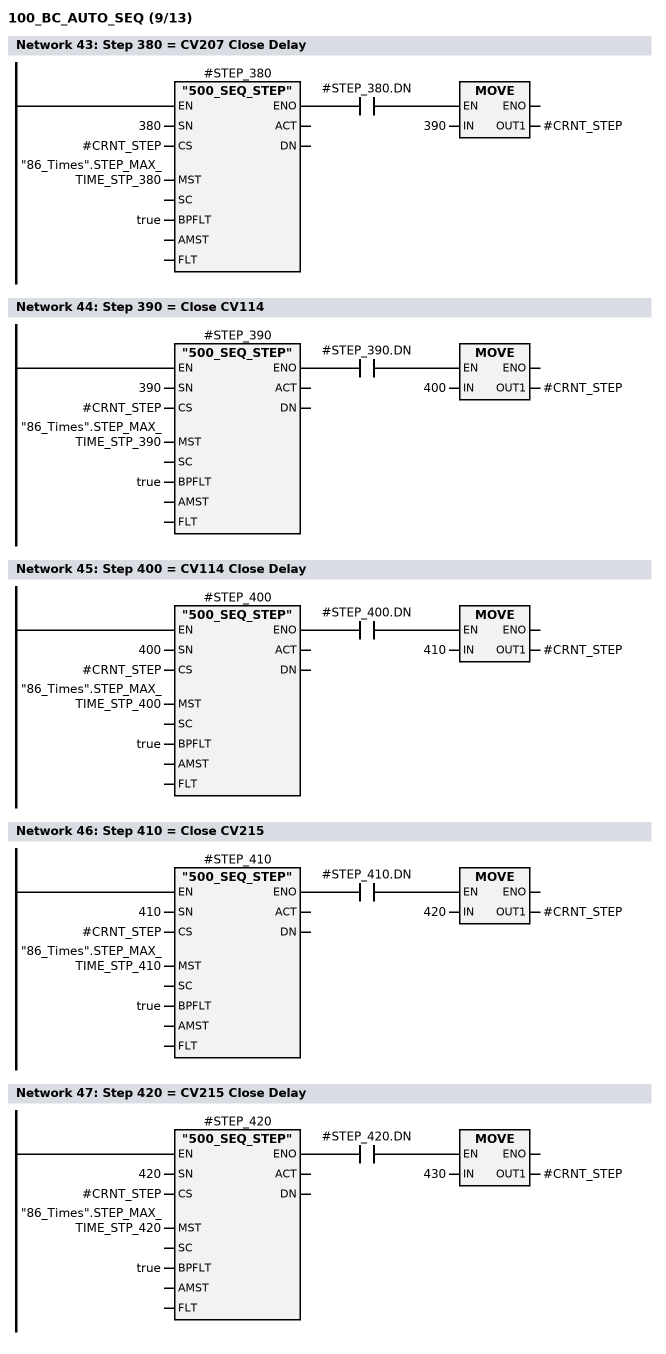
   RUNG wire#powerrail
      #STEP_380(SN := 380, CS := #CRNT_STEP, MST := "86_Times".STEP_MAX_TIME_STP_380, SC :=, BPFLT := true, AMST :=, FLT :=, ACT =>, DN =>)
      Contact( #STEP_380.DN )
      Move(in := 390, out1 => #CRNT_STEP)
   END_RUNG
   // the same network as SCL:
   #STEP_380(SN := 380, CS := #CRNT_STEP, MST := "86_Times".STEP_MAX_TIME_STP_380, BPFLT := true, ENO => #_w1);   // "500_SEQ_STEP"
   IF #_w1 AND #STEP_380.DN THEN #CRNT_STEP := 390; END_IF;
END_REGION

REGION Network 44: Step 390 = Close CV114
   RUNG wire#powerrail
      #STEP_390(SN := 390, CS := #CRNT_STEP, MST := "86_Times".STEP_MAX_TIME_STP_390, SC :=, BPFLT := true, AMST :=, FLT :=, ACT =>, DN =>)
      Contact( #STEP_390.DN )
      Move(in := 400, out1 => #CRNT_STEP)
   END_RUNG
   // the same network as SCL:
   #STEP_390(SN := 390, CS := #CRNT_STEP, MST := "86_Times".STEP_MAX_TIME_STP_390, BPFLT := true, ENO => #_w1);   // "500_SEQ_STEP"
   IF #_w1 AND #STEP_390.DN THEN #CRNT_STEP := 400; END_IF;
END_REGION

REGION Network 45: Step 400 = CV114 Close Delay
   RUNG wire#powerrail
      #STEP_400(SN := 400, CS := #CRNT_STEP, MST := "86_Times".STEP_MAX_TIME_STP_400, SC :=, BPFLT := true, AMST :=, FLT :=, ACT =>, DN =>)
      Contact( #STEP_400.DN )
      Move(in := 410, out1 => #CRNT_STEP)
   END_RUNG
   // the same network as SCL:
   #STEP_400(SN := 400, CS := #CRNT_STEP, MST := "86_Times".STEP_MAX_TIME_STP_400, BPFLT := true, ENO => #_w1);   // "500_SEQ_STEP"
   IF #_w1 AND #STEP_400.DN THEN #CRNT_STEP := 410; END_IF;
END_REGION

REGION Network 46: Step 410 = Close CV215
   RUNG wire#powerrail
      #STEP_410(SN := 410, CS := #CRNT_STEP, MST := "86_Times".STEP_MAX_TIME_STP_410, SC :=, BPFLT := true, AMST :=, FLT :=, ACT =>, DN =>)
      Contact( #STEP_410.DN )
      Move(in := 420, out1 => #CRNT_STEP)
   END_RUNG
   // the same network as SCL:
   #STEP_410(SN := 410, CS := #CRNT_STEP, MST := "86_Times".STEP_MAX_TIME_STP_410, BPFLT := true, ENO => #_w1);   // "500_SEQ_STEP"
   IF #_w1 AND #STEP_410.DN THEN #CRNT_STEP := 420; END_IF;
END_REGION

REGION Network 47: Step 420 = CV215 Close Delay
   RUNG wire#powerrail
      #STEP_420(SN := 420, CS := #CRNT_STEP, MST := "86_Times".STEP_MAX_TIME_STP_420, SC :=, BPFLT := true, AMST :=, FLT :=, ACT =>, DN =>)
      Contact( #STEP_420.DN )
      Move(in := 430, out1 => #CRNT_STEP)
   END_RUNG
   // the same network as SCL:
   #STEP_420(SN := 420, CS := #CRNT_STEP, MST := "86_Times".STEP_MAX_TIME_STP_420, BPFLT := true, ENO => #_w1);   // "500_SEQ_STEP"
   IF #_w1 AND #STEP_420.DN THEN #CRNT_STEP := 430; END_IF;
END_REGION

REGION Network 48: Step 430 = Close CV216
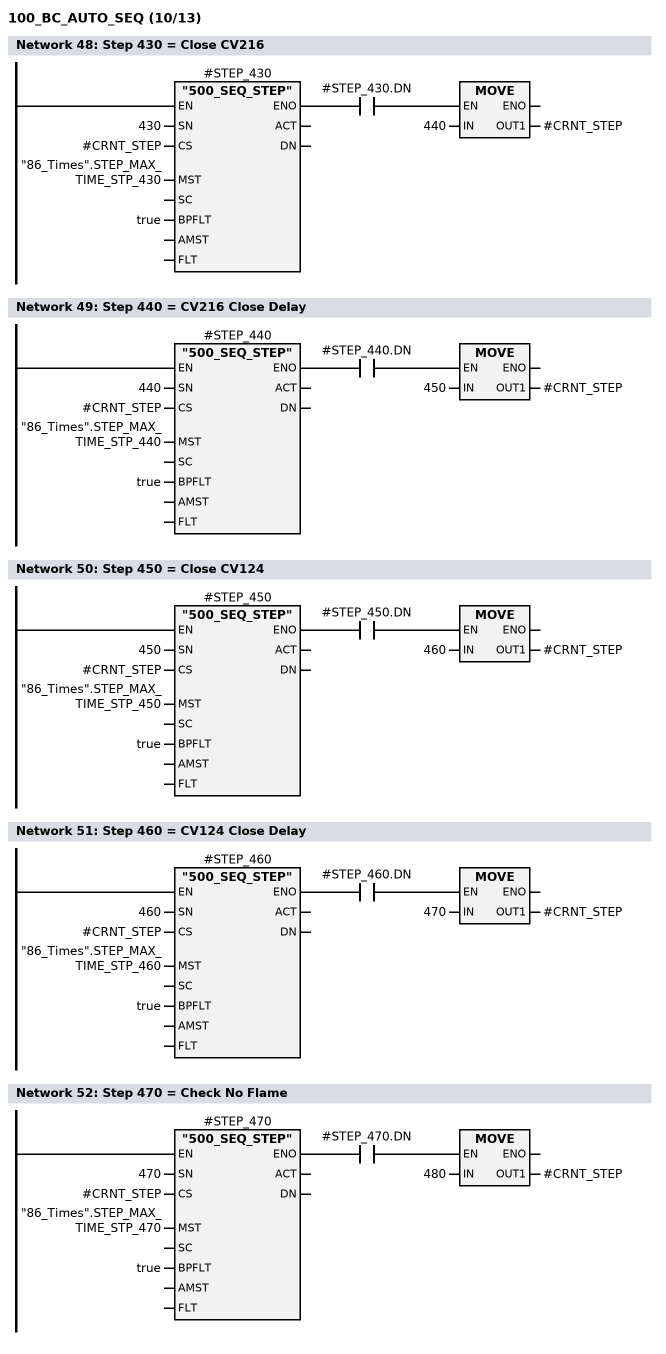
   RUNG wire#powerrail
      #STEP_430(SN := 430, CS := #CRNT_STEP, MST := "86_Times".STEP_MAX_TIME_STP_430, SC :=, BPFLT := true, AMST :=, FLT :=, ACT =>, DN =>)
      Contact( #STEP_430.DN )
      Move(in := 440, out1 => #CRNT_STEP)
   END_RUNG
   // the same network as SCL:
   #STEP_430(SN := 430, CS := #CRNT_STEP, MST := "86_Times".STEP_MAX_TIME_STP_430, BPFLT := true, ENO => #_w1);   // "500_SEQ_STEP"
   IF #_w1 AND #STEP_430.DN THEN #CRNT_STEP := 440; END_IF;
END_REGION

REGION Network 49: Step 440 = CV216 Close Delay
   RUNG wire#powerrail
      #STEP_440(SN := 440, CS := #CRNT_STEP, MST := "86_Times".STEP_MAX_TIME_STP_440, SC :=, BPFLT := true, AMST :=, FLT :=, ACT =>, DN =>)
      Contact( #STEP_440.DN )
      Move(in := 450, out1 => #CRNT_STEP)
   END_RUNG
   // the same network as SCL:
   #STEP_440(SN := 440, CS := #CRNT_STEP, MST := "86_Times".STEP_MAX_TIME_STP_440, BPFLT := true, ENO => #_w1);   // "500_SEQ_STEP"
   IF #_w1 AND #STEP_440.DN THEN #CRNT_STEP := 450; END_IF;
END_REGION

REGION Network 50: Step 450 = Close CV124
   RUNG wire#powerrail
      #STEP_450(SN := 450, CS := #CRNT_STEP, MST := "86_Times".STEP_MAX_TIME_STP_450, SC :=, BPFLT := true, AMST :=, FLT :=, ACT =>, DN =>)
      Contact( #STEP_450.DN )
      Move(in := 460, out1 => #CRNT_STEP)
   END_RUNG
   // the same network as SCL:
   #STEP_450(SN := 450, CS := #CRNT_STEP, MST := "86_Times".STEP_MAX_TIME_STP_450, BPFLT := true, ENO => #_w1);   // "500_SEQ_STEP"
   IF #_w1 AND #STEP_450.DN THEN #CRNT_STEP := 460; END_IF;
END_REGION

REGION Network 51: Step 460 = CV124 Close Delay
   RUNG wire#powerrail
      #STEP_460(SN := 460, CS := #CRNT_STEP, MST := "86_Times".STEP_MAX_TIME_STP_460, SC :=, BPFLT := true, AMST :=, FLT :=, ACT =>, DN =>)
      Contact( #STEP_460.DN )
      Move(in := 470, out1 => #CRNT_STEP)
   END_RUNG
   // the same network as SCL:
   #STEP_460(SN := 460, CS := #CRNT_STEP, MST := "86_Times".STEP_MAX_TIME_STP_460, BPFLT := true, ENO => #_w1);   // "500_SEQ_STEP"
   IF #_w1 AND #STEP_460.DN THEN #CRNT_STEP := 470; END_IF;
END_REGION

REGION Network 52: Step 470 = Check No Flame
   RUNG wire#powerrail
      #STEP_470(SN := 470, CS := #CRNT_STEP, MST := "86_Times".STEP_MAX_TIME_STP_470, SC :=, BPFLT := true, AMST :=, FLT :=, ACT =>, DN =>)
      Contact( #STEP_470.DN )
      Move(in := 480, out1 => #CRNT_STEP)
   END_RUNG
   // the same network as SCL:
   #STEP_470(SN := 470, CS := #CRNT_STEP, MST := "86_Times".STEP_MAX_TIME_STP_470, BPFLT := true, ENO => #_w1);   // "500_SEQ_STEP"
   IF #_w1 AND #STEP_470.DN THEN #CRNT_STEP := 480; END_IF;
END_REGION

REGION Network 53: Step 480 = Burn Stopped Confirmation To IGG
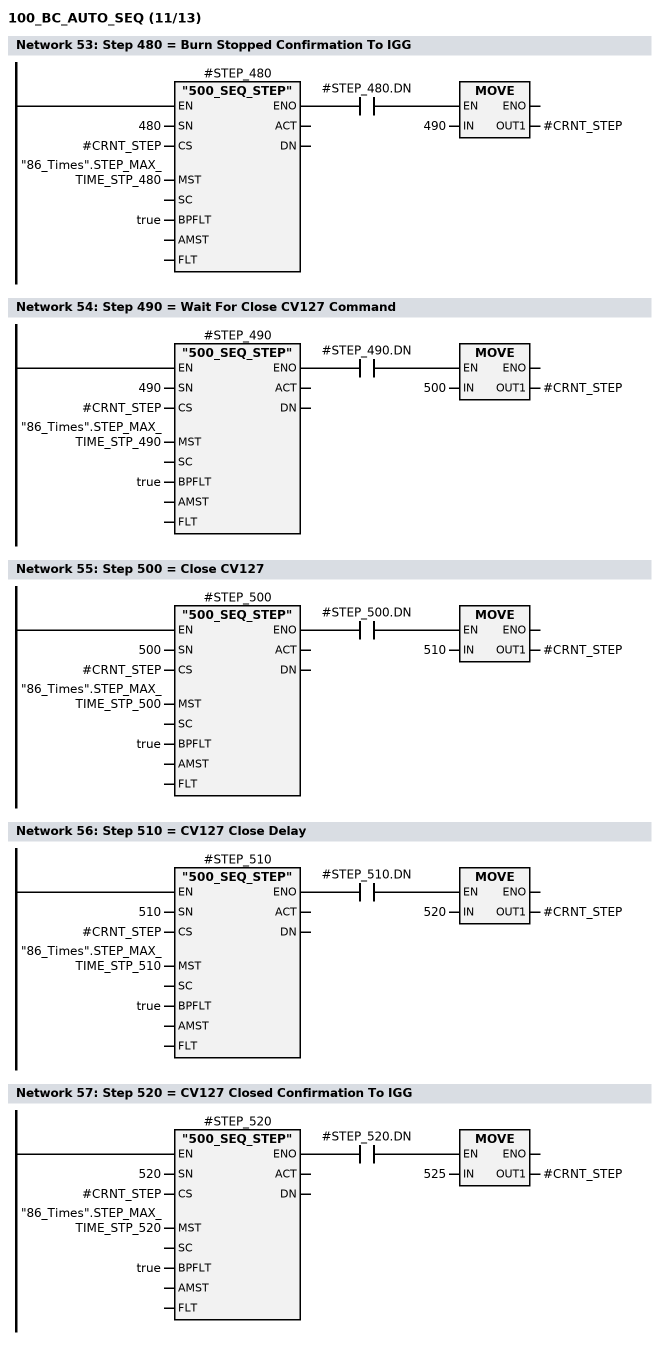
   RUNG wire#powerrail
      #STEP_480(SN := 480, CS := #CRNT_STEP, MST := "86_Times".STEP_MAX_TIME_STP_480, SC :=, BPFLT := true, AMST :=, FLT :=, ACT =>, DN =>)
      Contact( #STEP_480.DN )
      Move(in := 490, out1 => #CRNT_STEP)
   END_RUNG
   // the same network as SCL:
   #STEP_480(SN := 480, CS := #CRNT_STEP, MST := "86_Times".STEP_MAX_TIME_STP_480, BPFLT := true, ENO => #_w1);   // "500_SEQ_STEP"
   IF #_w1 AND #STEP_480.DN THEN #CRNT_STEP := 490; END_IF;
END_REGION

REGION Network 54: Step 490 = Wait For Close CV127 Command
   RUNG wire#powerrail
      #STEP_490(SN := 490, CS := #CRNT_STEP, MST := "86_Times".STEP_MAX_TIME_STP_490, SC :=, BPFLT := true, AMST :=, FLT :=, ACT =>, DN =>)
      Contact( #STEP_490.DN )
      Move(in := 500, out1 => #CRNT_STEP)
   END_RUNG
   // the same network as SCL:
   #STEP_490(SN := 490, CS := #CRNT_STEP, MST := "86_Times".STEP_MAX_TIME_STP_490, BPFLT := true, ENO => #_w1);   // "500_SEQ_STEP"
   IF #_w1 AND #STEP_490.DN THEN #CRNT_STEP := 500; END_IF;
END_REGION

REGION Network 55: Step 500 = Close CV127
   RUNG wire#powerrail
      #STEP_500(SN := 500, CS := #CRNT_STEP, MST := "86_Times".STEP_MAX_TIME_STP_500, SC :=, BPFLT := true, AMST :=, FLT :=, ACT =>, DN =>)
      Contact( #STEP_500.DN )
      Move(in := 510, out1 => #CRNT_STEP)
   END_RUNG
   // the same network as SCL:
   #STEP_500(SN := 500, CS := #CRNT_STEP, MST := "86_Times".STEP_MAX_TIME_STP_500, BPFLT := true, ENO => #_w1);   // "500_SEQ_STEP"
   IF #_w1 AND #STEP_500.DN THEN #CRNT_STEP := 510; END_IF;
END_REGION

REGION Network 56: Step 510 = CV127 Close Delay
   RUNG wire#powerrail
      #STEP_510(SN := 510, CS := #CRNT_STEP, MST := "86_Times".STEP_MAX_TIME_STP_510, SC :=, BPFLT := true, AMST :=, FLT :=, ACT =>, DN =>)
      Contact( #STEP_510.DN )
      Move(in := 520, out1 => #CRNT_STEP)
   END_RUNG
   // the same network as SCL:
   #STEP_510(SN := 510, CS := #CRNT_STEP, MST := "86_Times".STEP_MAX_TIME_STP_510, BPFLT := true, ENO => #_w1);   // "500_SEQ_STEP"
   IF #_w1 AND #STEP_510.DN THEN #CRNT_STEP := 520; END_IF;
END_REGION

REGION Network 57: Step 520 = CV127 Closed Confirmation To IGG
   RUNG wire#powerrail
      #STEP_520(SN := 520, CS := #CRNT_STEP, MST := "86_Times".STEP_MAX_TIME_STP_520, SC :=, BPFLT := true, AMST :=, FLT :=, ACT =>, DN =>)
      Contact( #STEP_520.DN )
      Move(in := 525, out1 => #CRNT_STEP)
   END_RUNG
   // the same network as SCL:
   #STEP_520(SN := 520, CS := #CRNT_STEP, MST := "86_Times".STEP_MAX_TIME_STP_520, BPFLT := true, ENO => #_w1);   // "500_SEQ_STEP"
   IF #_w1 AND #STEP_520.DN THEN #CRNT_STEP := 525; END_IF;
END_REGION

REGION Network 58: Step 525 = Wait For Close CV203 Command
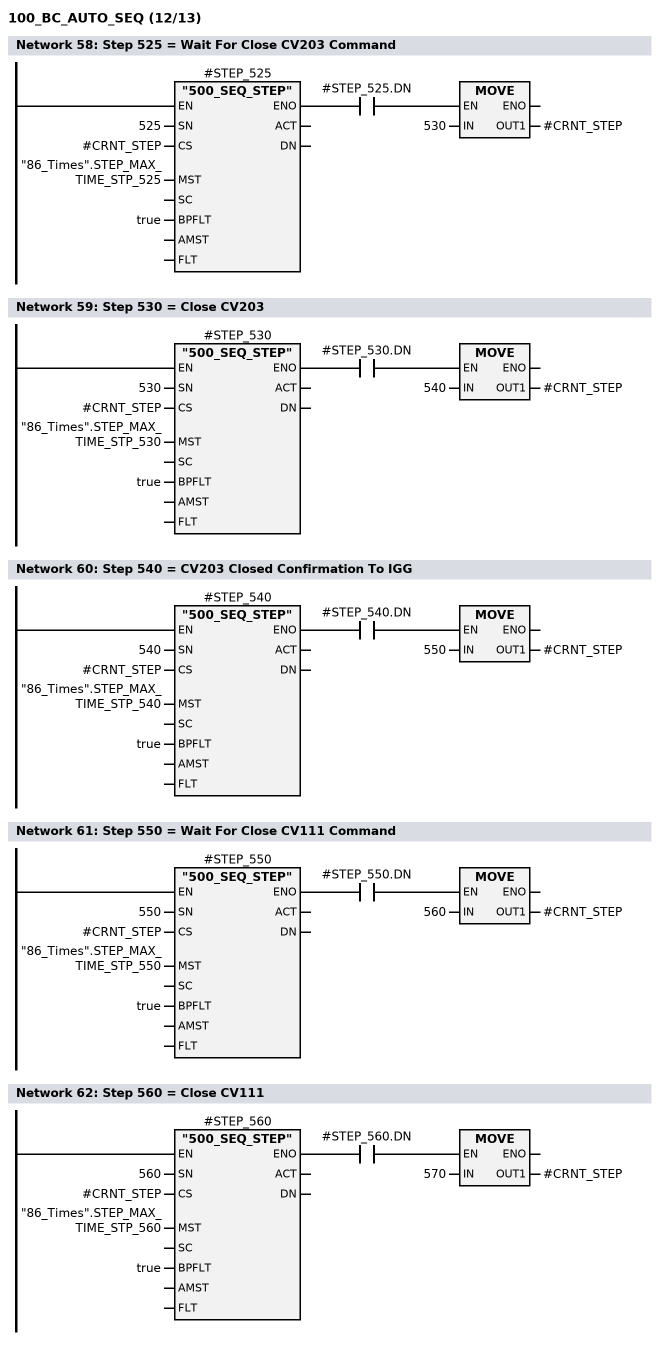
   RUNG wire#powerrail
      #STEP_525(SN := 525, CS := #CRNT_STEP, MST := "86_Times".STEP_MAX_TIME_STP_525, SC :=, BPFLT := true, AMST :=, FLT :=, ACT =>, DN =>)
      Contact( #STEP_525.DN )
      Move(in := 530, out1 => #CRNT_STEP)
   END_RUNG
   // the same network as SCL:
   #STEP_525(SN := 525, CS := #CRNT_STEP, MST := "86_Times".STEP_MAX_TIME_STP_525, BPFLT := true, ENO => #_w1);   // "500_SEQ_STEP"
   IF #_w1 AND #STEP_525.DN THEN #CRNT_STEP := 530; END_IF;
END_REGION

REGION Network 59: Step 530 = Close CV203
   RUNG wire#powerrail
      #STEP_530(SN := 530, CS := #CRNT_STEP, MST := "86_Times".STEP_MAX_TIME_STP_530, SC :=, BPFLT := true, AMST :=, FLT :=, ACT =>, DN =>)
      Contact( #STEP_530.DN )
      Move(in := 540, out1 => #CRNT_STEP)
   END_RUNG
   // the same network as SCL:
   #STEP_530(SN := 530, CS := #CRNT_STEP, MST := "86_Times".STEP_MAX_TIME_STP_530, BPFLT := true, ENO => #_w1);   // "500_SEQ_STEP"
   IF #_w1 AND #STEP_530.DN THEN #CRNT_STEP := 540; END_IF;
END_REGION

REGION Network 60: Step 540 = CV203 Closed Confirmation To IGG
   RUNG wire#powerrail
      #STEP_540(SN := 540, CS := #CRNT_STEP, MST := "86_Times".STEP_MAX_TIME_STP_540, SC :=, BPFLT := true, AMST :=, FLT :=, ACT =>, DN =>)
      Contact( #STEP_540.DN )
      Move(in := 550, out1 => #CRNT_STEP)
   END_RUNG
   // the same network as SCL:
   #STEP_540(SN := 540, CS := #CRNT_STEP, MST := "86_Times".STEP_MAX_TIME_STP_540, BPFLT := true, ENO => #_w1);   // "500_SEQ_STEP"
   IF #_w1 AND #STEP_540.DN THEN #CRNT_STEP := 550; END_IF;
END_REGION

REGION Network 61: Step 550 = Wait For Close CV111 Command
   RUNG wire#powerrail
      #STEP_550(SN := 550, CS := #CRNT_STEP, MST := "86_Times".STEP_MAX_TIME_STP_550, SC :=, BPFLT := true, AMST :=, FLT :=, ACT =>, DN =>)
      Contact( #STEP_550.DN )
      Move(in := 560, out1 => #CRNT_STEP)
   END_RUNG
   // the same network as SCL:
   #STEP_550(SN := 550, CS := #CRNT_STEP, MST := "86_Times".STEP_MAX_TIME_STP_550, BPFLT := true, ENO => #_w1);   // "500_SEQ_STEP"
   IF #_w1 AND #STEP_550.DN THEN #CRNT_STEP := 560; END_IF;
END_REGION

REGION Network 62: Step 560 = Close CV111
   RUNG wire#powerrail
      #STEP_560(SN := 560, CS := #CRNT_STEP, MST := "86_Times".STEP_MAX_TIME_STP_560, SC :=, BPFLT := true, AMST :=, FLT :=, ACT =>, DN =>)
      Contact( #STEP_560.DN )
      Move(in := 570, out1 => #CRNT_STEP)
   END_RUNG
   // the same network as SCL:
   #STEP_560(SN := 560, CS := #CRNT_STEP, MST := "86_Times".STEP_MAX_TIME_STP_560, BPFLT := true, ENO => #_w1);   // "500_SEQ_STEP"
   IF #_w1 AND #STEP_560.DN THEN #CRNT_STEP := 570; END_IF;
END_REGION

REGION Network 63: Step 570 = Shutdown Done Status To IGG
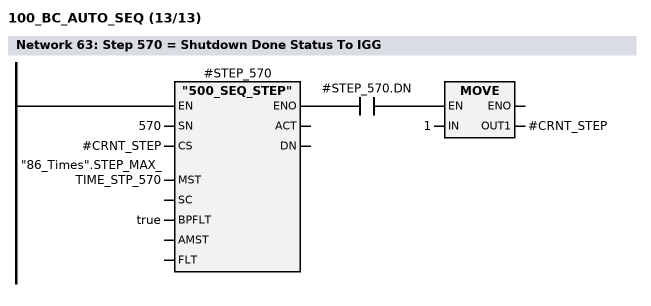
   RUNG wire#powerrail
      #STEP_570(SN := 570, CS := #CRNT_STEP, MST := "86_Times".STEP_MAX_TIME_STP_570, SC :=, BPFLT := true, AMST :=, FLT :=, ACT =>, DN =>)
      Contact( #STEP_570.DN )
      Move(in := 1, out1 => #CRNT_STEP)
   END_RUNG
   // the same network as SCL:
   #STEP_570(SN := 570, CS := #CRNT_STEP, MST := "86_Times".STEP_MAX_TIME_STP_570, BPFLT := true, ENO => #_w1);   // "500_SEQ_STEP"
   IF #_w1 AND #STEP_570.DN THEN #CRNT_STEP := 1; END_IF;
END_REGION
END_FUNCTION_BLOCK

FUNCTION_BLOCK "102_Pilot_Burner"   // FB102, LAD
TITLE = Pilot Burner Control
{ S7_Optimized_Access := 'TRUE' }
AUTHOR : JRS
VERSION : 0.1
// For the control of the pilot burner ignition and burn
   VAR_INPUT
      RUN : Bool;   // Runs the block
      FLM_DET : Bool;   // Flame detected
      FLM_FAIL_DLY : Time;
      IGNTR_DLY : Time;   // Igniter delay time
      IGNTR_MAX_RT : Time;   // Igniter maximum run time
      FV1_DLY : Time;   // Fuel valve 1 delay time
      FV2_3W_DLY : Time;   // 3 Way fuel valve 2 delay time
      FD_DLY : Time;   // Flame detection delay time
      FD_SCAN_TIME : Time;   // Flame detection scan time
      FD_VRFCTN_TIME : Time;   // Flame verification time
      MAX_SEQ_TIME : Time;   // Maximum sequence run time
      IGNTR_PWR_OK : Bool;   // Igniter power ok
      FDU_PWR_OK : Bool;   // Flame detection unit power ok
      FDU_OK : Bool;   // Flame detection health ok
      RST : Bool;   // Reset bit
   END_VAR
   VAR_OUTPUT
      RUN_IGNTR : Bool;   // Run igniter
      OPN_FV1 : Bool;   // Open fuel valve 1
      OPN_3W_FV2 : Bool;   // Open 3 way fuel valve 2
      DN_OK : Bool;   // Successful ignition
      IAC : Int;   // Ignition atttempt count
      FAILED : Bool;   // Ignition failed
      FLT : Bool;   // Fault bit
   END_VAR
   VAR_IN_OUT
      RUNNING : Bool;   // Sequence running
   END_VAR
   VAR
      INTO_RUN_EDGE : Bool;   // Edge detection
      OUT_OF_RUN_EDGE : Bool;   // Edge detection
      LOOK_NEG_EDGE : Bool;   // Stop looking edge
      INTO_S20 : Bool;   // Into step 20
      INTO_S20_EDGE : Bool;   // Into step 20 edge
      RST_FLG : Bool;   // Reset flag
      LOOKING : Bool;   // Looking for flame
      STATE : Int;   // State value for sequencing
      IAC_VAL : Int;   // Ignition attempt count value
      IGNTR_TMR : TOF_TIME;   // Igniter maximum run time
      FD_SCN_TMR : TOF_TIME;   // Flame detection scan timer
      IGNTR_DLY_TMR : TON_TIME;   // Igniter delay timer
      IGNTR_STP_TMR : TON_TIME;   // Igniter stop timer
      FV1_DLY_TMR : TON_TIME;   // Fuel valve 1 delay timer
      FV2_DLY_TMR : TON_TIME;   // Fuel valve 2 delay timer
      FD_DLY_TMR : TON_TIME;   // Flame detection delay timer
      FD_VRFCTN_TMR : TON_TIME;   // Flame verification timer
      MAX_SEQ_TMR : TON_TIME;   // Maximum sequence run timer
      FV1_CLS_DLY_TMR : TON_TIME;   // Fuel valve 1 close delay timer
      FV2_CLS_DLY_TMR : TON_TIME;   // Fuel valve 2 close delay timer
      FLM_FAIL_TON : TON_TIME;
      "FD_VRFCTN_TMR II" : TON_TIME;
   END_VAR
   VAR_TEMP   // added for the SCL form of the ladder/FBD networks
      _w1 : Bool;
   END_VAR
BEGIN

REGION Network 1: Running
   // For running status detection
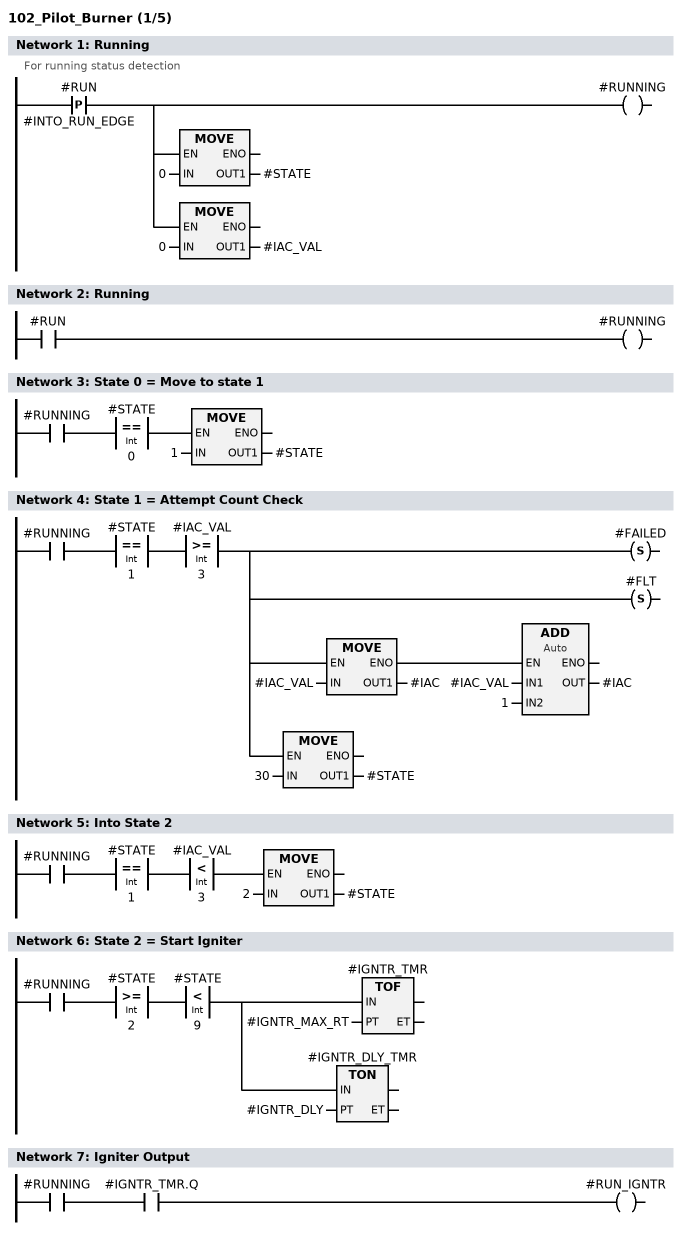
   RUNG wire#powerrail
      P_Contact(operand := #RUN, bit := #INTO_RUN_EDGE)
      wire#w1
      Coil( #RUNNING )
   END_RUNG
   RUNG wire#w1
      Move(in := 0, out1 => #STATE)
   END_RUNG
   RUNG wire#w1
      Move(in := 0, out1 => #IAC_VAL)
   END_RUNG
   // the same network as SCL:
   #_w1 := #RUN AND NOT #INTO_RUN_EDGE;   // rising edge of #RUN
   #INTO_RUN_EDGE := #RUN;
   #RUNNING := #_w1;
   IF #_w1 THEN
       #STATE := 0;
       #IAC_VAL := 0;
   END_IF;
END_REGION

REGION Network 2: Running
   RUNG wire#powerrail
      Contact( #RUN )
      Coil( #RUNNING )
   END_RUNG
   // the same network as SCL:
   #RUNNING := #RUN;
END_REGION

REGION Network 3: State 0 = Move to state 1
   RUNG wire#powerrail
      Contact( #RUNNING )
      { S7_Templates := "SrcType := Int" } EQ_Contact(in1 := #STATE, in2 := 0)
      Move(in := 1, out1 => #STATE)
   END_RUNG
   // the same network as SCL:
   IF #RUNNING AND (#STATE = 0) THEN #STATE := 1; END_IF;
END_REGION

REGION Network 4: State 1 = Attempt Count Check
   RUNG wire#powerrail
      Contact( #RUNNING )
      { S7_Templates := "SrcType := Int" } EQ_Contact(in1 := #STATE, in2 := 1)
      { S7_Templates := "SrcType := Int" } GE_Contact(in1 := #IAC_VAL, in2 := 3)
      wire#w1
      S_Coil( #FAILED )
   END_RUNG
   RUNG wire#w1
      S_Coil( #FLT )
   END_RUNG
   RUNG wire#w1
      Move(in := #IAC_VAL, out1 => #IAC)
      Add(in1 := #IAC_VAL, in2 := 1, out => #IAC)
   END_RUNG
   RUNG wire#w1
      Move(in := 30, out1 => #STATE)
   END_RUNG
   // the same network as SCL:
   IF #RUNNING AND (#STATE = 1) AND (#IAC_VAL >= 3) THEN
       #FAILED := TRUE;
       #FLT := TRUE;
       #IAC := #IAC_VAL;
       #IAC := #IAC_VAL + 1;
       #STATE := 30;
   END_IF;
END_REGION

REGION Network 5: Into State 2
   RUNG wire#powerrail
      Contact( #RUNNING )
      { S7_Templates := "SrcType := Int" } EQ_Contact(in1 := #STATE, in2 := 1)
      { S7_Templates := "SrcType := Int" } LT_Contact(in1 := #IAC_VAL, in2 := 3)
      Move(in := 2, out1 => #STATE)
   END_RUNG
   // the same network as SCL:
   IF #RUNNING AND (#STATE = 1) AND (#IAC_VAL < 3) THEN #STATE := 2; END_IF;
END_REGION

REGION Network 6: State 2 = Start Igniter
   #_w1 := #RUNNING AND (#STATE >= 2) AND (#STATE < 9);
   #IGNTR_TMR(IN := #_w1, PT := #IGNTR_MAX_RT);   // TOF
   #IGNTR_DLY_TMR(IN := #_w1, PT := #IGNTR_DLY);   // TON
END_REGION

REGION Network 7: Igniter Output
   RUNG wire#powerrail
      Contact( #RUNNING )
      Contact( #IGNTR_TMR.Q )
      Coil( #RUN_IGNTR )
   END_RUNG
   // the same network as SCL:
   #RUN_IGNTR := #RUNNING AND #IGNTR_TMR.Q;
END_REGION

REGION Network 8: Into State 3
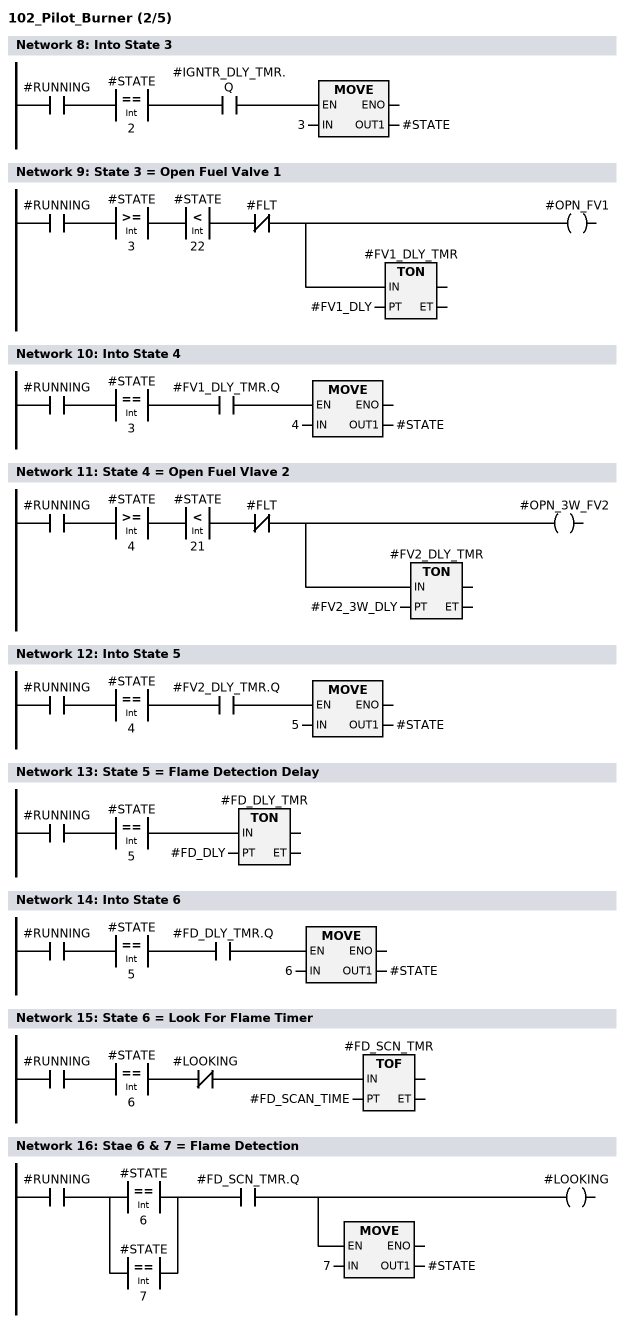
   RUNG wire#powerrail
      Contact( #RUNNING )
      { S7_Templates := "SrcType := Int" } EQ_Contact(in1 := #STATE, in2 := 2)
      Contact( #IGNTR_DLY_TMR.Q )
      Move(in := 3, out1 => #STATE)
   END_RUNG
   // the same network as SCL:
   IF #RUNNING AND (#STATE = 2) AND #IGNTR_DLY_TMR.Q THEN #STATE := 3; END_IF;
END_REGION

REGION Network 9: State 3 = Open Fuel Valve 1
   #OPN_FV1 := #RUNNING AND (#STATE >= 3) AND (#STATE < 22) AND NOT #FLT;
   #FV1_DLY_TMR(IN := #OPN_FV1, PT := #FV1_DLY);   // TON
END_REGION

REGION Network 10: Into State 4
   RUNG wire#powerrail
      Contact( #RUNNING )
      { S7_Templates := "SrcType := Int" } EQ_Contact(in1 := #STATE, in2 := 3)
      Contact( #FV1_DLY_TMR.Q )
      Move(in := 4, out1 => #STATE)
   END_RUNG
   // the same network as SCL:
   IF #RUNNING AND (#STATE = 3) AND #FV1_DLY_TMR.Q THEN #STATE := 4; END_IF;
END_REGION

REGION Network 11: State 4 = Open Fuel Vlave 2
   #OPN_3W_FV2 := #RUNNING AND (#STATE >= 4) AND (#STATE < 21) AND NOT #FLT;
   #FV2_DLY_TMR(IN := #OPN_3W_FV2, PT := #FV2_3W_DLY);   // TON
END_REGION

REGION Network 12: Into State 5
   RUNG wire#powerrail
      Contact( #RUNNING )
      { S7_Templates := "SrcType := Int" } EQ_Contact(in1 := #STATE, in2 := 4)
      Contact( #FV2_DLY_TMR.Q )
      Move(in := 5, out1 => #STATE)
   END_RUNG
   // the same network as SCL:
   IF #RUNNING AND (#STATE = 4) AND #FV2_DLY_TMR.Q THEN #STATE := 5; END_IF;
END_REGION

REGION Network 13: State 5 = Flame Detection Delay
   #FD_DLY_TMR(IN := #RUNNING AND (#STATE = 5), PT := #FD_DLY);   // TON
END_REGION

REGION Network 14: Into State 6
   RUNG wire#powerrail
      Contact( #RUNNING )
      { S7_Templates := "SrcType := Int" } EQ_Contact(in1 := #STATE, in2 := 5)
      Contact( #FD_DLY_TMR.Q )
      Move(in := 6, out1 => #STATE)
   END_RUNG
   // the same network as SCL:
   IF #RUNNING AND (#STATE = 5) AND #FD_DLY_TMR.Q THEN #STATE := 6; END_IF;
END_REGION

REGION Network 15: State 6 = Look For Flame Timer
   #FD_SCN_TMR(IN := #RUNNING AND (#STATE = 6) AND NOT #LOOKING, PT := #FD_SCAN_TIME);   // TOF
END_REGION

REGION Network 16: Stae 6 & 7 = Flame Detection
   RUNG wire#powerrail
      Contact( #RUNNING )
      wire#w1
      { S7_Templates := "SrcType := Int" } EQ_Contact(in1 := #STATE, in2 := 6)
      wire#w2
      Contact( #FD_SCN_TMR.Q )
      wire#w3
      Coil( #LOOKING )
   END_RUNG
   RUNG wire#w1
      { S7_Templates := "SrcType := Int" } EQ_Contact(in1 := #STATE, in2 := 7)
   END_RUNG wire#w2
   RUNG wire#w3
      Move(in := 7, out1 => #STATE)
   END_RUNG
   // the same network as SCL:
   #LOOKING := #RUNNING AND ((#STATE = 6) OR (#STATE = 7)) AND #FD_SCN_TMR.Q;
   IF #LOOKING THEN #STATE := 7; END_IF;
END_REGION

REGION Network 17: Flame Detection = Move To Step 8
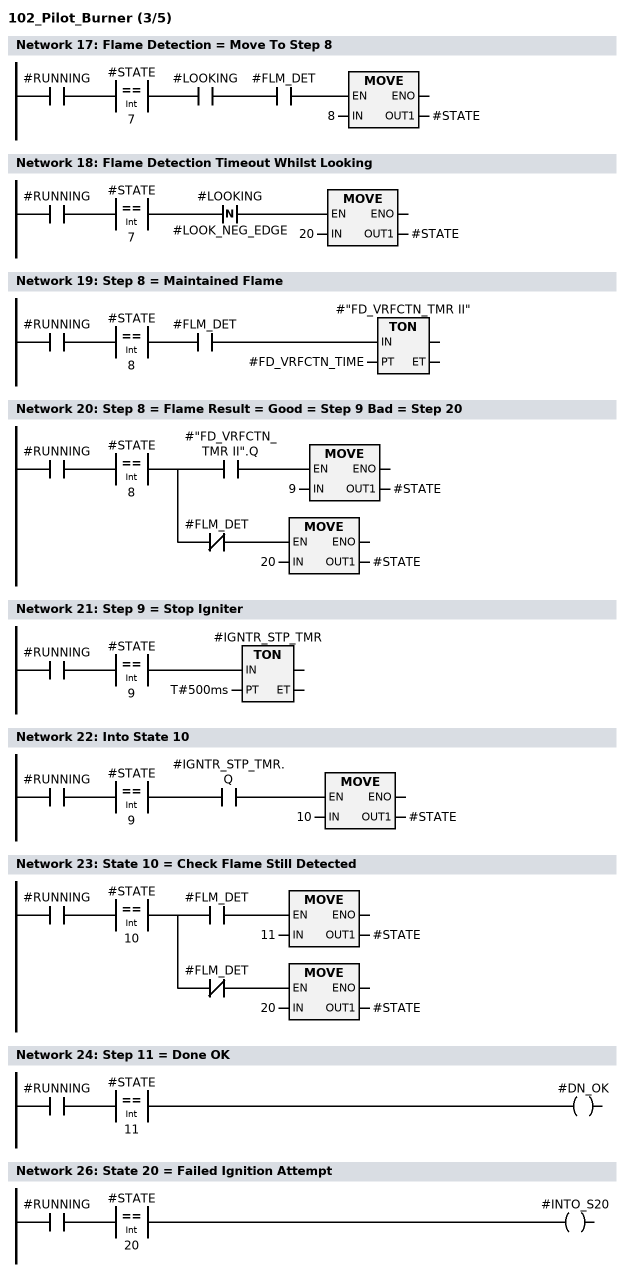
   RUNG wire#powerrail
      Contact( #RUNNING )
      { S7_Templates := "SrcType := Int" } EQ_Contact(in1 := #STATE, in2 := 7)
      Contact( #LOOKING )
      Contact( #FLM_DET )
      Move(in := 8, out1 => #STATE)
   END_RUNG
   // the same network as SCL:
   IF #RUNNING AND (#STATE = 7) AND #LOOKING AND #FLM_DET THEN #STATE := 8; END_IF;
END_REGION

REGION Network 18: Flame Detection Timeout Whilst Looking
   RUNG wire#powerrail
      Contact( #RUNNING )
      { S7_Templates := "SrcType := Int" } EQ_Contact(in1 := #STATE, in2 := 7)
      N_Contact(operand := #LOOKING, bit := #LOOK_NEG_EDGE)
      Move(in := 20, out1 => #STATE)
   END_RUNG
   // the same network as SCL:
   #_w1 := #RUNNING AND (#STATE = 7) AND NOT #LOOKING AND #LOOK_NEG_EDGE;   // falling edge of #LOOKING
   #LOOK_NEG_EDGE := #LOOKING;
   IF #_w1 THEN #STATE := 20; END_IF;
END_REGION

REGION Network 19: Step 8 = Maintained Flame
   #"FD_VRFCTN_TMR II"(IN := #RUNNING AND (#STATE = 8) AND #FLM_DET, PT := #FD_VRFCTN_TIME);   // TON
END_REGION

REGION Network 20: Step 8 = Flame Result = Good = Step 9 Bad = Step 20
   RUNG wire#powerrail
      Contact( #RUNNING )
      { S7_Templates := "SrcType := Int" } EQ_Contact(in1 := #STATE, in2 := 8)
      wire#w1
      Contact( #"FD_VRFCTN_TMR II".Q )
      Move(in := 9, out1 => #STATE)
   END_RUNG
   RUNG wire#w1
      I_Contact( #FLM_DET )
      Move(in := 20, out1 => #STATE)
   END_RUNG
   // the same network as SCL:
   #_w1 := #RUNNING AND (#STATE = 8);
   IF #_w1 AND #"FD_VRFCTN_TMR II".Q THEN #STATE := 9; END_IF;
   IF #_w1 AND NOT #FLM_DET THEN #STATE := 20; END_IF;
END_REGION

REGION Network 21: Step 9 = Stop Igniter
   #IGNTR_STP_TMR(IN := #RUNNING AND (#STATE = 9), PT := T#500ms);   // TON
END_REGION

REGION Network 22: Into State 10
   RUNG wire#powerrail
      Contact( #RUNNING )
      { S7_Templates := "SrcType := Int" } EQ_Contact(in1 := #STATE, in2 := 9)
      Contact( #IGNTR_STP_TMR.Q )
      Move(in := 10, out1 => #STATE)
   END_RUNG
   // the same network as SCL:
   IF #RUNNING AND (#STATE = 9) AND #IGNTR_STP_TMR.Q THEN #STATE := 10; END_IF;
END_REGION

REGION Network 23: State 10 = Check Flame Still Detected
   RUNG wire#powerrail
      Contact( #RUNNING )
      { S7_Templates := "SrcType := Int" } EQ_Contact(in1 := #STATE, in2 := 10)
      wire#w1
      Contact( #FLM_DET )
      Move(in := 11, out1 => #STATE)
   END_RUNG
   RUNG wire#w1
      I_Contact( #FLM_DET )
      Move(in := 20, out1 => #STATE)
   END_RUNG
   // the same network as SCL:
   #_w1 := #RUNNING AND (#STATE = 10);
   IF #_w1 AND #FLM_DET THEN #STATE := 11; END_IF;
   IF #_w1 AND NOT #FLM_DET THEN #STATE := 20; END_IF;
END_REGION

REGION Network 24: Step 11 = Done OK
   RUNG wire#powerrail
      Contact( #RUNNING )
      { S7_Templates := "SrcType := Int" } EQ_Contact(in1 := #STATE, in2 := 11)
      Coil( #DN_OK )
   END_RUNG
   // the same network as SCL:
   #DN_OK := #RUNNING AND (#STATE = 11);
END_REGION

REGION Network 26: State 20 = Failed Ignition Attempt
   RUNG wire#powerrail
      Contact( #RUNNING )
      { S7_Templates := "SrcType := Int" } EQ_Contact(in1 := #STATE, in2 := 20)
      Coil( #INTO_S20 )
   END_RUNG
   // the same network as SCL:
   #INTO_S20 := #RUNNING AND (#STATE = 20);
END_REGION